// TIA Portal project "SMS-ENLAB-01-003-1501-001-PLC_V13_SP1_2_V17" (V17) (continued)
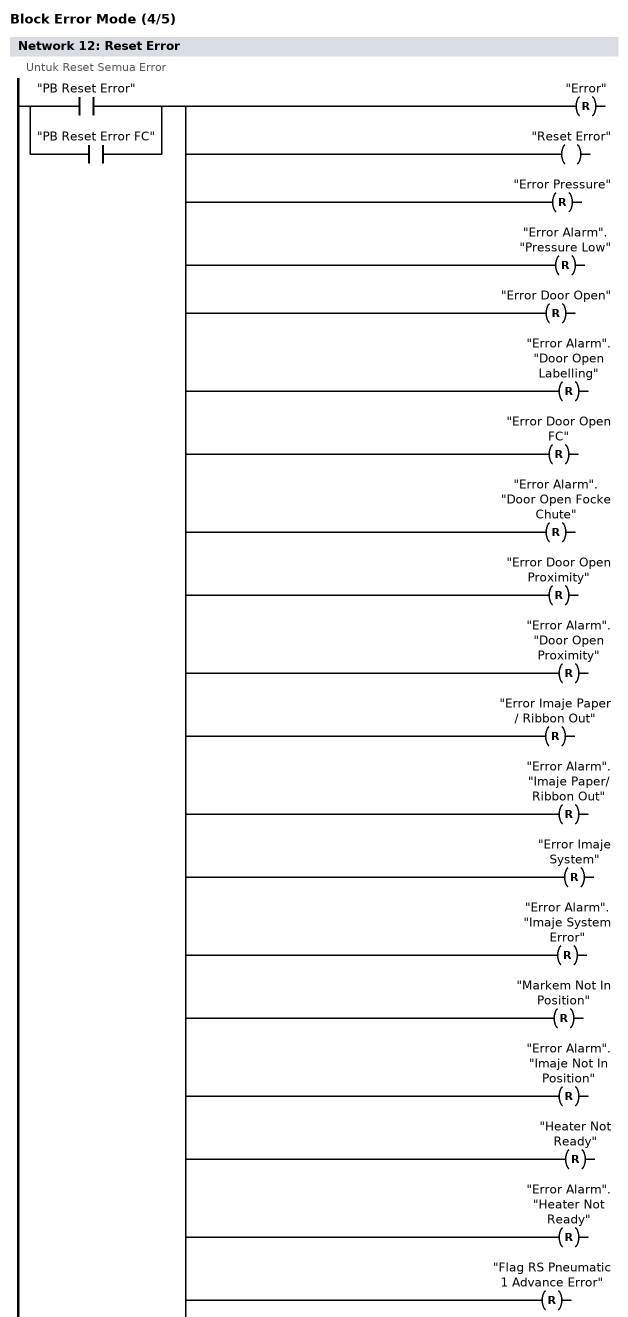
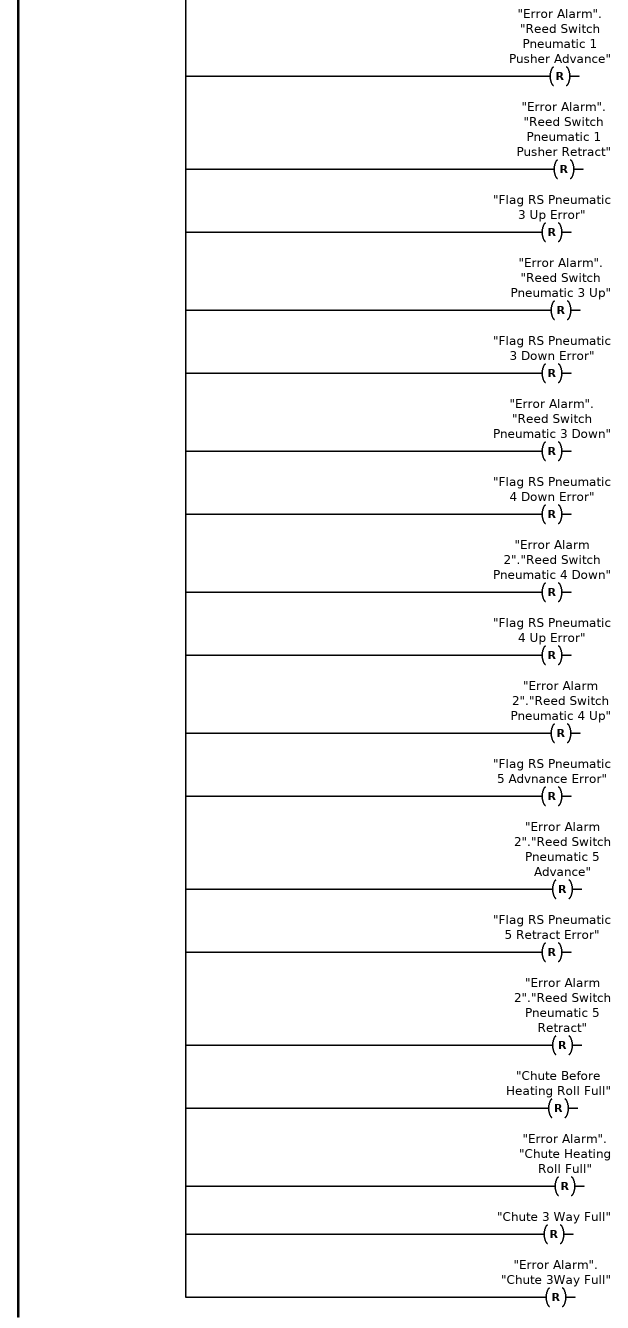
   RUNG wire#powerrail
      Contact( "PB Reset Error" )
      wire#w1
      R_Coil( "Error" )
   END_RUNG
   RUNG wire#powerrail
      Contact( "PB Reset Error FC" )
   END_RUNG wire#w1
   RUNG wire#w1
      Coil( "Reset Error" )
   END_RUNG
   RUNG wire#w1
      R_Coil( "Error Pressure" )
   END_RUNG
   RUNG wire#w1
      R_Coil( "Error Alarm"."Pressure Low" )
   END_RUNG
   RUNG wire#w1
      R_Coil( "Error Door Open" )
   END_RUNG
   RUNG wire#w1
      R_Coil( "Error Alarm"."Door Open Labelling" )
   END_RUNG
   RUNG wire#w1
      R_Coil( "Error Door Open FC" )
   END_RUNG
   RUNG wire#w1
      R_Coil( "Error Alarm"."Door Open Focke Chute" )
   END_RUNG
   RUNG wire#w1
      R_Coil( "Error Door Open Proximity" )
   END_RUNG
   RUNG wire#w1
      R_Coil( "Error Alarm"."Door Open Proximity" )
   END_RUNG
   RUNG wire#w1
      R_Coil( "Error Imaje Paper / Ribbon Out" )
   END_RUNG
   RUNG wire#w1
      R_Coil( "Error Alarm"."Imaje Paper/Ribbon Out" )
   END_RUNG
   RUNG wire#w1
      R_Coil( "Error Imaje System" )
   END_RUNG
   RUNG wire#w1
      R_Coil( "Error Alarm"."Imaje System Error" )
   END_RUNG
   RUNG wire#w1
      R_Coil( "Markem Not In Position" )
   END_RUNG
   RUNG wire#w1
      R_Coil( "Error Alarm"."Imaje Not In Position" )
   END_RUNG
   RUNG wire#w1
      R_Coil( "Heater Not Ready" )
   END_RUNG
   RUNG wire#w1
      R_Coil( "Error Alarm"."Heater Not Ready" )
   END_RUNG
   RUNG wire#w1
      R_Coil( "Flag RS Pneumatic 1 Advance Error" )
   END_RUNG
   RUNG wire#w1
      R_Coil( "Error Alarm"."Reed Switch Pneumatic 1 Pusher Advance" )
   END_RUNG
   RUNG wire#w1
      R_Coil( "Error Alarm"."Reed Switch Pneumatic 1 Pusher Retract" )
   END_RUNG
   RUNG wire#w1
      R_Coil( "Flag RS Pneumatic 3 Up Error" )
   END_RUNG
   RUNG wire#w1
      R_Coil( "Error Alarm"."Reed Switch Pneumatic 3 Up" )
   END_RUNG
   RUNG wire#w1
      R_Coil( "Flag RS Pneumatic 3 Down Error" )
   END_RUNG
   RUNG wire#w1
      R_Coil( "Error Alarm"."Reed Switch Pneumatic 3 Down" )
   END_RUNG
   RUNG wire#w1
      R_Coil( "Flag RS Pneumatic 4 Down Error" )
   END_RUNG
   RUNG wire#w1
      R_Coil( "Error Alarm 2"."Reed Switch Pneumatic 4 Down" )
   END_RUNG
   RUNG wire#w1
      R_Coil( "Flag RS Pneumatic 4 Up Error" )
   END_RUNG
   RUNG wire#w1
      R_Coil( "Error Alarm 2"."Reed Switch Pneumatic 4 Up" )
   END_RUNG
   RUNG wire#w1
      R_Coil( "Flag RS Pneumatic 5 Advnance Error" )
   END_RUNG
   RUNG wire#w1
      R_Coil( "Error Alarm 2"."Reed Switch Pneumatic 5 Advance" )
   END_RUNG
   RUNG wire#w1
      R_Coil( "Flag RS Pneumatic 5 Retract Error" )
   END_RUNG
   RUNG wire#w1
      R_Coil( "Error Alarm 2"."Reed Switch Pneumatic 5 Retract" )
   END_RUNG
   RUNG wire#w1
      R_Coil( "Chute Before Heating Roll Full" )
   END_RUNG
   RUNG wire#w1
      R_Coil( "Error Alarm"."Chute Heating Roll Full" )
   END_RUNG
   RUNG wire#w1
      R_Coil( "Chute 3 Way Full" )
   END_RUNG
   RUNG wire#w1
      R_Coil( "Error Alarm"."Chute 3Way Full" )
   END_RUNG
   // the same network as SCL:
   #_w1 := "PB Reset Error" OR "PB Reset Error FC";
   IF #_w1 THEN "Error" := FALSE; END_IF;
   "Reset Error" := #_w1;
   IF #_w1 THEN
       "Error Pressure" := FALSE;
       "Error Alarm"."Pressure Low" := FALSE;
       "Error Door Open" := FALSE;
       "Error Alarm"."Door Open Labelling" := FALSE;
       "Error Door Open FC" := FALSE;
       "Error Alarm"."Door Open Focke Chute" := FALSE;
       "Error Door Open Proximity" := FALSE;
       "Error Alarm"."Door Open Proximity" := FALSE;
       "Error Imaje Paper / Ribbon Out" := FALSE;
       "Error Alarm"."Imaje Paper/Ribbon Out" := FALSE;
       "Error Imaje System" := FALSE;
       "Error Alarm"."Imaje System Error" := FALSE;
       "Markem Not In Position" := FALSE;
       "Error Alarm"."Imaje Not In Position" := FALSE;
       "Heater Not Ready" := FALSE;
       "Error Alarm"."Heater Not Ready" := FALSE;
       "Flag RS Pneumatic 1 Advance Error" := FALSE;
       "Error Alarm"."Reed Switch Pneumatic 1 Pusher Advance" := FALSE;
       "Error Alarm"."Reed Switch Pneumatic 1 Pusher Retract" := FALSE;
       "Flag RS Pneumatic 3 Up Error" := FALSE;
       "Error Alarm"."Reed Switch Pneumatic 3 Up" := FALSE;
       "Flag RS Pneumatic 3 Down Error" := FALSE;
       "Error Alarm"."Reed Switch Pneumatic 3 Down" := FALSE;
       "Flag RS Pneumatic 4 Down Error" := FALSE;
       "Error Alarm 2"."Reed Switch Pneumatic 4 Down" := FALSE;
       "Flag RS Pneumatic 4 Up Error" := FALSE;
       "Error Alarm 2"."Reed Switch Pneumatic 4 Up" := FALSE;
       "Flag RS Pneumatic 5 Advnance Error" := FALSE;
       "Error Alarm 2"."Reed Switch Pneumatic 5 Advance" := FALSE;
       "Flag RS Pneumatic 5 Retract Error" := FALSE;
       "Error Alarm 2"."Reed Switch Pneumatic 5 Retract" := FALSE;
       "Chute Before Heating Roll Full" := FALSE;
       "Error Alarm"."Chute Heating Roll Full" := FALSE;
       "Chute 3 Way Full" := FALSE;
       "Error Alarm"."Chute 3Way Full" := FALSE;
   END_IF;
END_REGION

REGION Network 13: Enable Flow to Reject
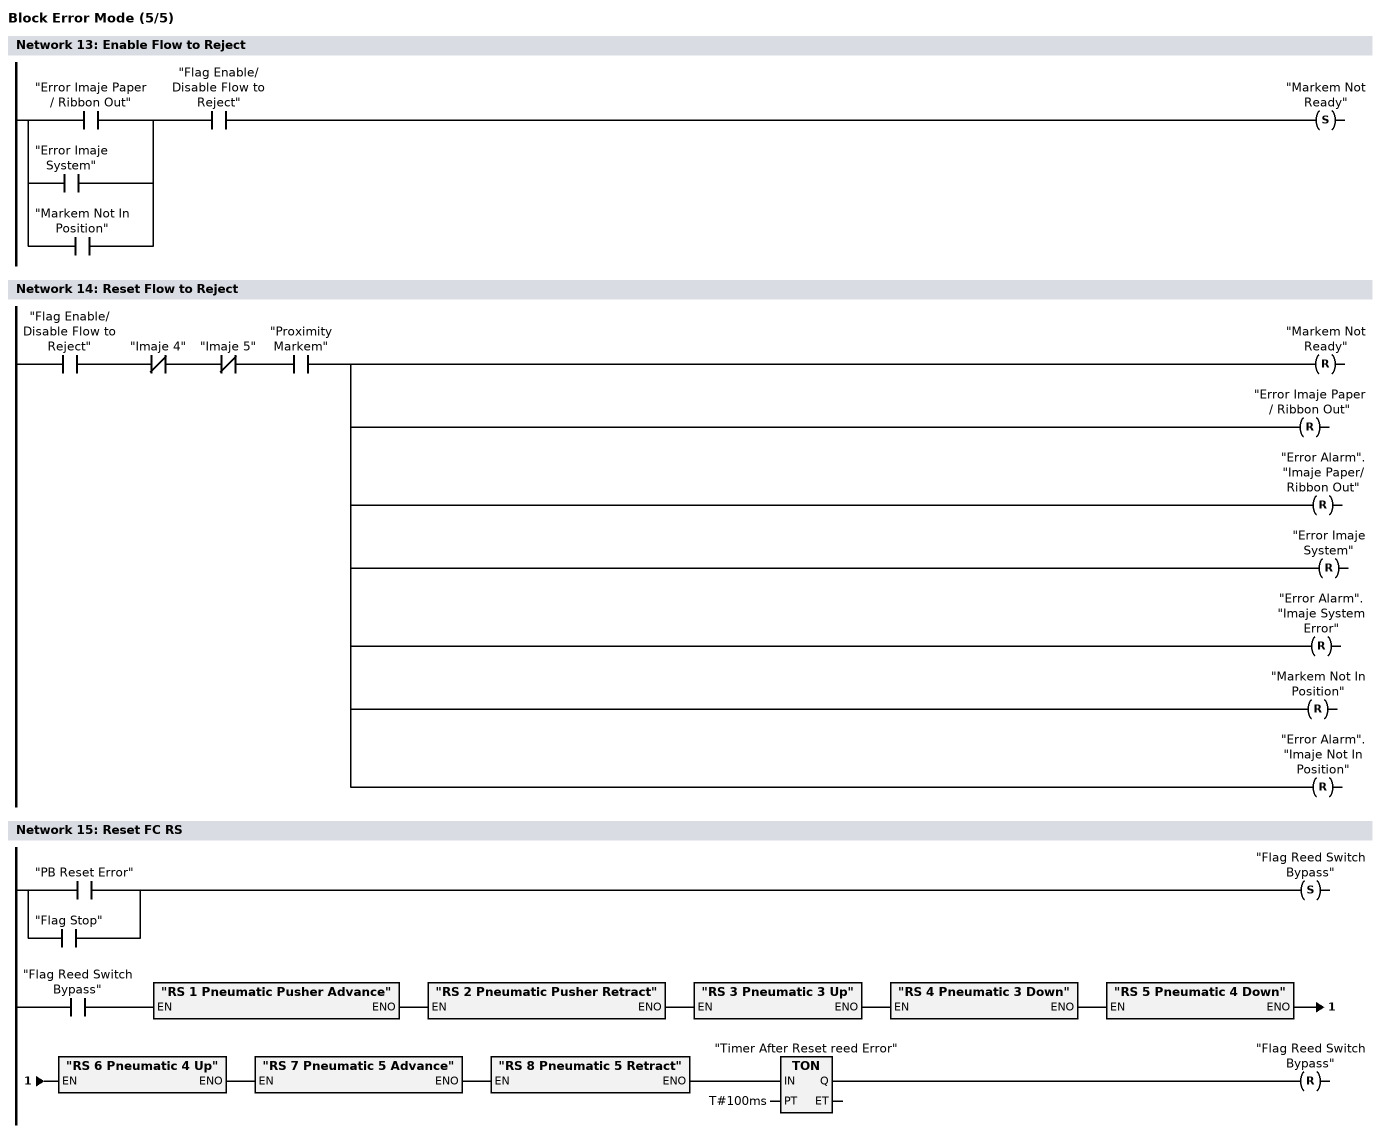
   RUNG wire#powerrail
      Contact( "Error Imaje Paper / Ribbon Out" )
      wire#w1
      Contact( "Flag Enable/Disable Flow to Reject" )
      S_Coil( "Markem Not Ready" )
   END_RUNG
   RUNG wire#powerrail
      Contact( "Error Imaje System" )
   END_RUNG wire#w1
   RUNG wire#powerrail
      Contact( "Markem Not In Position" )
   END_RUNG wire#w1
   // the same network as SCL:
   IF ("Error Imaje Paper / Ribbon Out" OR "Error Imaje System" OR "Markem Not In Position") AND "Flag Enable/Disable Flow to Reject" THEN
       "Markem Not Ready" := TRUE;
   END_IF;
END_REGION

REGION Network 14: Reset Flow to Reject
   RUNG wire#powerrail
      Contact( "Flag Enable/Disable Flow to Reject" )
      I_Contact( "Imaje 4" )
      I_Contact( "Imaje 5" )
      Contact( "Proximity Markem" )
      wire#w1
      R_Coil( "Markem Not Ready" )
   END_RUNG
   RUNG wire#w1
      R_Coil( "Error Imaje Paper / Ribbon Out" )
   END_RUNG
   RUNG wire#w1
      R_Coil( "Error Alarm"."Imaje Paper/Ribbon Out" )
   END_RUNG
   RUNG wire#w1
      R_Coil( "Error Imaje System" )
   END_RUNG
   RUNG wire#w1
      R_Coil( "Error Alarm"."Imaje System Error" )
   END_RUNG
   RUNG wire#w1
      R_Coil( "Markem Not In Position" )
   END_RUNG
   RUNG wire#w1
      R_Coil( "Error Alarm"."Imaje Not In Position" )
   END_RUNG
   // the same network as SCL:
   IF "Flag Enable/Disable Flow to Reject" AND NOT "Imaje 4" AND NOT "Imaje 5" AND "Proximity Markem" THEN
       "Markem Not Ready" := FALSE;
       "Error Imaje Paper / Ribbon Out" := FALSE;
       "Error Alarm"."Imaje Paper/Ribbon Out" := FALSE;
       "Error Imaje System" := FALSE;
       "Error Alarm"."Imaje System Error" := FALSE;
       "Markem Not In Position" := FALSE;
       "Error Alarm"."Imaje Not In Position" := FALSE;
   END_IF;
END_REGION

REGION Network 15: Reset FC RS
   IF "PB Reset Error" OR "Flag Stop" THEN "Flag Reed Switch Bypass" := TRUE; END_IF;
   "RS 1 Pneumatic Pusher Advance"(EN := "Flag Reed Switch Bypass", ENO => #_w1);
   "RS 2 Pneumatic Pusher Retract"(EN := #_w1, ENO => #_w2);
   "RS 3 Pneumatic 3 Up"(EN := #_w2, ENO => #_w3);
   "RS 4 Pneumatic 3 Down"(EN := #_w3, ENO => #_w4);
   "RS 5 Pneumatic 4 Down"(EN := #_w4, ENO => #_w5);
   "RS 6 Pneumatic 4 Up"(EN := #_w5, ENO => #_w6);
   "RS 7 Pneumatic 5 Advance"(EN := #_w6, ENO => #_w7);
   "RS 8 Pneumatic 5 Retract"(EN := #_w7, ENO => #_w8);
   "Timer After Reset reed Error".TON(IN := #_w8, PT := T#100ms);
   IF "Timer After Reset reed Error".Q THEN "Flag Reed Switch Bypass" := FALSE; END_IF;
END_REGION
END_FUNCTION_BLOCK

FUNCTION_BLOCK "Block Test Mode"   // FB2, LAD
{ S7_Optimized_Access := 'TRUE' }
VERSION : 0.1
BEGIN

REGION Network 1: Set Motor Conveyor
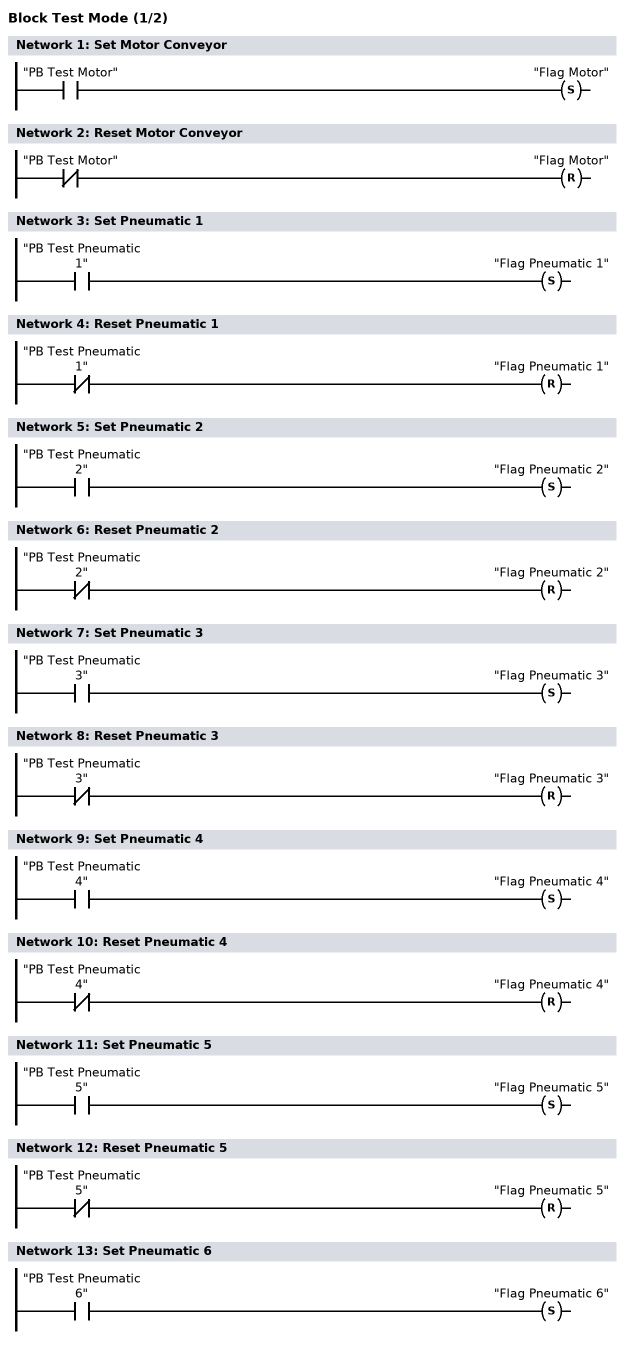
   RUNG wire#powerrail
      Contact( "PB Test Motor" )
      S_Coil( "Flag Motor" )
   END_RUNG
   // the same network as SCL:
   IF "PB Test Motor" THEN "Flag Motor" := TRUE; END_IF;
END_REGION

REGION Network 2: Reset Motor Conveyor
   RUNG wire#powerrail
      I_Contact( "PB Test Motor" )
      R_Coil( "Flag Motor" )
   END_RUNG
   // the same network as SCL:
   IF NOT "PB Test Motor" THEN "Flag Motor" := FALSE; END_IF;
END_REGION

REGION Network 3: Set Pneumatic 1
   RUNG wire#powerrail
      Contact( "PB Test Pneumatic 1" )
      S_Coil( "Flag Pneumatic 1" )
   END_RUNG
   // the same network as SCL:
   IF "PB Test Pneumatic 1" THEN "Flag Pneumatic 1" := TRUE; END_IF;
END_REGION

REGION Network 4: Reset Pneumatic 1
   RUNG wire#powerrail
      I_Contact( "PB Test Pneumatic 1" )
      R_Coil( "Flag Pneumatic 1" )
   END_RUNG
   // the same network as SCL:
   IF NOT "PB Test Pneumatic 1" THEN "Flag Pneumatic 1" := FALSE; END_IF;
END_REGION

REGION Network 5: Set Pneumatic 2
   RUNG wire#powerrail
      Contact( "PB Test Pneumatic 2" )
      S_Coil( "Flag Pneumatic 2" )
   END_RUNG
   // the same network as SCL:
   IF "PB Test Pneumatic 2" THEN "Flag Pneumatic 2" := TRUE; END_IF;
END_REGION

REGION Network 6: Reset Pneumatic 2
   RUNG wire#powerrail
      I_Contact( "PB Test Pneumatic 2" )
      R_Coil( "Flag Pneumatic 2" )
   END_RUNG
   // the same network as SCL:
   IF NOT "PB Test Pneumatic 2" THEN "Flag Pneumatic 2" := FALSE; END_IF;
END_REGION

REGION Network 7: Set Pneumatic 3
   RUNG wire#powerrail
      Contact( "PB Test Pneumatic 3" )
      S_Coil( "Flag Pneumatic 3" )
   END_RUNG
   // the same network as SCL:
   IF "PB Test Pneumatic 3" THEN "Flag Pneumatic 3" := TRUE; END_IF;
END_REGION

REGION Network 8: Reset Pneumatic 3
   RUNG wire#powerrail
      I_Contact( "PB Test Pneumatic 3" )
      R_Coil( "Flag Pneumatic 3" )
   END_RUNG
   // the same network as SCL:
   IF NOT "PB Test Pneumatic 3" THEN "Flag Pneumatic 3" := FALSE; END_IF;
END_REGION

REGION Network 9: Set Pneumatic 4
   RUNG wire#powerrail
      Contact( "PB Test Pneumatic 4" )
      S_Coil( "Flag Pneumatic 4" )
   END_RUNG
   // the same network as SCL:
   IF "PB Test Pneumatic 4" THEN "Flag Pneumatic 4" := TRUE; END_IF;
END_REGION

REGION Network 10: Reset Pneumatic 4
   RUNG wire#powerrail
      I_Contact( "PB Test Pneumatic 4" )
      R_Coil( "Flag Pneumatic 4" )
   END_RUNG
   // the same network as SCL:
   IF NOT "PB Test Pneumatic 4" THEN "Flag Pneumatic 4" := FALSE; END_IF;
END_REGION

REGION Network 11: Set Pneumatic 5
   RUNG wire#powerrail
      Contact( "PB Test Pneumatic 5" )
      S_Coil( "Flag Pneumatic 5" )
   END_RUNG
   // the same network as SCL:
   IF "PB Test Pneumatic 5" THEN "Flag Pneumatic 5" := TRUE; END_IF;
END_REGION

REGION Network 12: Reset Pneumatic 5
   RUNG wire#powerrail
      I_Contact( "PB Test Pneumatic 5" )
      R_Coil( "Flag Pneumatic 5" )
   END_RUNG
   // the same network as SCL:
   IF NOT "PB Test Pneumatic 5" THEN "Flag Pneumatic 5" := FALSE; END_IF;
END_REGION

REGION Network 13: Set Pneumatic 6
   RUNG wire#powerrail
      Contact( "PB Test Pneumatic 6" )
      S_Coil( "Flag Pneumatic 6" )
   END_RUNG
   // the same network as SCL:
   IF "PB Test Pneumatic 6" THEN "Flag Pneumatic 6" := TRUE; END_IF;
END_REGION

REGION Network 14: Reset Pneumatic 6
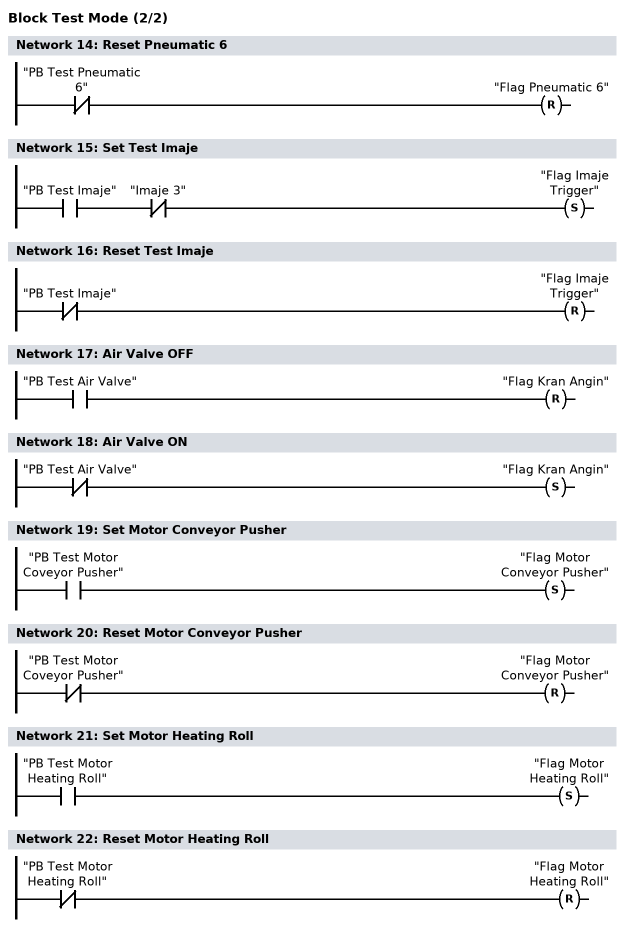
   RUNG wire#powerrail
      I_Contact( "PB Test Pneumatic 6" )
      R_Coil( "Flag Pneumatic 6" )
   END_RUNG
   // the same network as SCL:
   IF NOT "PB Test Pneumatic 6" THEN "Flag Pneumatic 6" := FALSE; END_IF;
END_REGION

REGION Network 15: Set Test Imaje
   RUNG wire#powerrail
      Contact( "PB Test Imaje" )
      I_Contact( "Imaje 3" )
      S_Coil( "Flag Imaje Trigger" )
   END_RUNG
   // the same network as SCL:
   IF "PB Test Imaje" AND NOT "Imaje 3" THEN "Flag Imaje Trigger" := TRUE; END_IF;
END_REGION

REGION Network 16: Reset Test Imaje
   RUNG wire#powerrail
      I_Contact( "PB Test Imaje" )
      R_Coil( "Flag Imaje Trigger" )
   END_RUNG
   // the same network as SCL:
   IF NOT "PB Test Imaje" THEN "Flag Imaje Trigger" := FALSE; END_IF;
END_REGION

REGION Network 17: Air Valve OFF
   RUNG wire#powerrail
      Contact( "PB Test Air Valve" )
      R_Coil( "Flag Kran Angin" )
   END_RUNG
   // the same network as SCL:
   IF "PB Test Air Valve" THEN "Flag Kran Angin" := FALSE; END_IF;
END_REGION

REGION Network 18: Air Valve ON
   RUNG wire#powerrail
      I_Contact( "PB Test Air Valve" )
      S_Coil( "Flag Kran Angin" )
   END_RUNG
   // the same network as SCL:
   IF NOT "PB Test Air Valve" THEN "Flag Kran Angin" := TRUE; END_IF;
END_REGION

REGION Network 19: Set Motor Conveyor Pusher
   RUNG wire#powerrail
      Contact( "PB Test Motor Coveyor Pusher" )
      S_Coil( "Flag Motor Conveyor Pusher" )
   END_RUNG
   // the same network as SCL:
   IF "PB Test Motor Coveyor Pusher" THEN "Flag Motor Conveyor Pusher" := TRUE; END_IF;
END_REGION

REGION Network 20: Reset Motor Conveyor Pusher
   RUNG wire#powerrail
      I_Contact( "PB Test Motor Coveyor Pusher" )
      R_Coil( "Flag Motor Conveyor Pusher" )
   END_RUNG
   // the same network as SCL:
   IF NOT "PB Test Motor Coveyor Pusher" THEN "Flag Motor Conveyor Pusher" := FALSE; END_IF;
END_REGION

REGION Network 21: Set Motor Heating Roll
   RUNG wire#powerrail
      Contact( "PB Test Motor Heating Roll" )
      S_Coil( "Flag Motor Heating Roll" )
   END_RUNG
   // the same network as SCL:
   IF "PB Test Motor Heating Roll" THEN "Flag Motor Heating Roll" := TRUE; END_IF;
END_REGION

REGION Network 22: Reset Motor Heating Roll
   RUNG wire#powerrail
      I_Contact( "PB Test Motor Heating Roll" )
      R_Coil( "Flag Motor Heating Roll" )
   END_RUNG
   // the same network as SCL:
   IF NOT "PB Test Motor Heating Roll" THEN "Flag Motor Heating Roll" := FALSE; END_IF;
END_REGION
END_FUNCTION_BLOCK

FUNCTION_BLOCK "Block Output"   // FB3, LAD
{ S7_Optimized_Access := 'TRUE' }
VERSION : 0.1
BEGIN

REGION Network 1: Red Light Tower
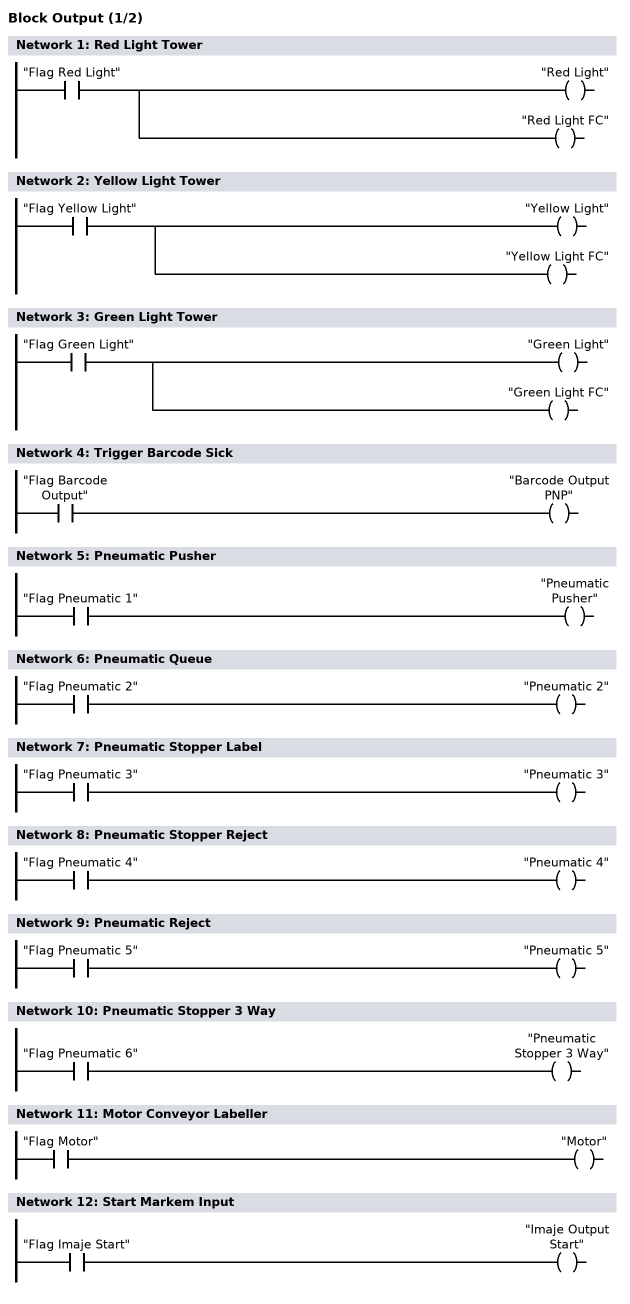
   RUNG wire#powerrail
      Contact( "Flag Red Light" )
      wire#w1
      Coil( "Red Light" )
   END_RUNG
   RUNG wire#w1
      Coil( "Red Light FC" )
   END_RUNG
   // the same network as SCL:
   "Red Light" := "Flag Red Light";
   "Red Light FC" := "Flag Red Light";
END_REGION

REGION Network 2: Yellow Light Tower
   RUNG wire#powerrail
      Contact( "Flag Yellow Light" )
      wire#w1
      Coil( "Yellow Light" )
   END_RUNG
   RUNG wire#w1
      Coil( "Yellow Light FC" )
   END_RUNG
   // the same network as SCL:
   "Yellow Light" := "Flag Yellow Light";
   "Yellow Light FC" := "Flag Yellow Light";
END_REGION

REGION Network 3: Green Light Tower
   RUNG wire#powerrail
      Contact( "Flag Green Light" )
      wire#w1
      Coil( "Green Light" )
   END_RUNG
   RUNG wire#w1
      Coil( "Green Light FC" )
   END_RUNG
   // the same network as SCL:
   "Green Light" := "Flag Green Light";
   "Green Light FC" := "Flag Green Light";
END_REGION

REGION Network 4: Trigger Barcode Sick
   RUNG wire#powerrail
      Contact( "Flag Barcode Output" )
      Coil( "Barcode Output PNP" )
   END_RUNG
   // the same network as SCL:
   "Barcode Output PNP" := "Flag Barcode Output";
END_REGION

REGION Network 5: Pneumatic Pusher
   RUNG wire#powerrail
      Contact( "Flag Pneumatic 1" )
      Coil( "Pneumatic Pusher" )
   END_RUNG
   // the same network as SCL:
   "Pneumatic Pusher" := "Flag Pneumatic 1";
END_REGION

REGION Network 6: Pneumatic Queue
   RUNG wire#powerrail
      Contact( "Flag Pneumatic 2" )
      Coil( "Pneumatic 2" )
   END_RUNG
   // the same network as SCL:
   "Pneumatic 2" := "Flag Pneumatic 2";
END_REGION

REGION Network 7: Pneumatic Stopper Label
   RUNG wire#powerrail
      Contact( "Flag Pneumatic 3" )
      Coil( "Pneumatic 3" )
   END_RUNG
   // the same network as SCL:
   "Pneumatic 3" := "Flag Pneumatic 3";
END_REGION

REGION Network 8: Pneumatic Stopper Reject
   RUNG wire#powerrail
      Contact( "Flag Pneumatic 4" )
      Coil( "Pneumatic 4" )
   END_RUNG
   // the same network as SCL:
   "Pneumatic 4" := "Flag Pneumatic 4";
END_REGION

REGION Network 9: Pneumatic Reject
   RUNG wire#powerrail
      Contact( "Flag Pneumatic 5" )
      Coil( "Pneumatic 5" )
   END_RUNG
   // the same network as SCL:
   "Pneumatic 5" := "Flag Pneumatic 5";
END_REGION

REGION Network 10: Pneumatic Stopper 3 Way
   RUNG wire#powerrail
      Contact( "Flag Pneumatic 6" )
      Coil( "Pneumatic Stopper 3 Way" )
   END_RUNG
   // the same network as SCL:
   "Pneumatic Stopper 3 Way" := "Flag Pneumatic 6";
END_REGION

REGION Network 11: Motor Conveyor Labeller
   RUNG wire#powerrail
      Contact( "Flag Motor" )
      Coil( "Motor" )
   END_RUNG
   // the same network as SCL:
   "Motor" := "Flag Motor";
END_REGION

REGION Network 12: Start Markem Input
   RUNG wire#powerrail
      Contact( "Flag Imaje Start" )
      Coil( "Imaje Output Start" )
   END_RUNG
   // the same network as SCL:
   "Imaje Output Start" := "Flag Imaje Start";
END_REGION

REGION Network 13: Pause Markem Input
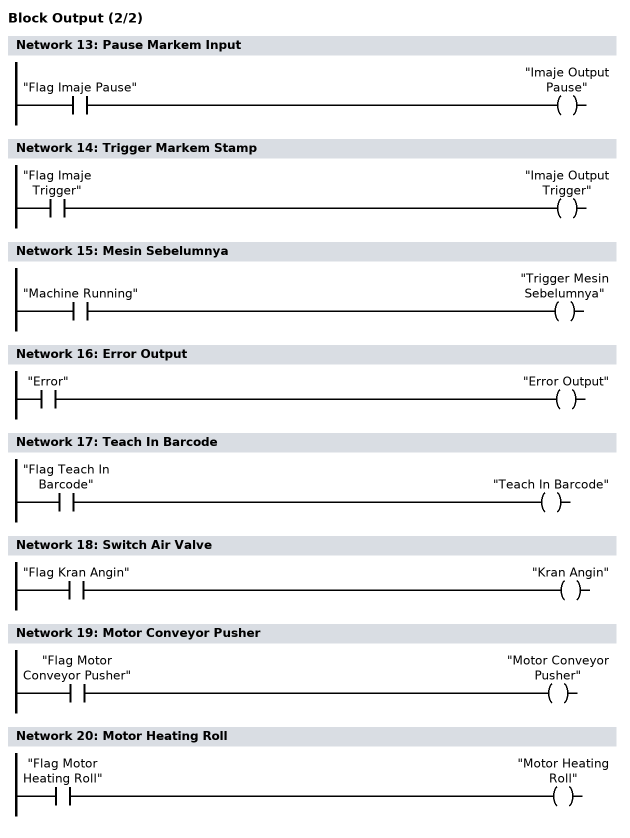
   RUNG wire#powerrail
      Contact( "Flag Imaje Pause" )
      Coil( "Imaje Output Pause" )
   END_RUNG
   // the same network as SCL:
   "Imaje Output Pause" := "Flag Imaje Pause";
END_REGION

REGION Network 14: Trigger Markem Stamp
   RUNG wire#powerrail
      Contact( "Flag Imaje Trigger" )
      Coil( "Imaje Output Trigger" )
   END_RUNG
   // the same network as SCL:
   "Imaje Output Trigger" := "Flag Imaje Trigger";
END_REGION

REGION Network 15: Mesin Sebelumnya
   RUNG wire#powerrail
      Contact( "Machine Running" )
      Coil( "Trigger Mesin Sebelumnya" )
   END_RUNG
   // the same network as SCL:
   "Trigger Mesin Sebelumnya" := "Machine Running";
END_REGION

REGION Network 16: Error Output
   RUNG wire#powerrail
      Contact( "Error" )
      Coil( "Error Output" )
   END_RUNG
   // the same network as SCL:
   "Error Output" := "Error";
END_REGION

REGION Network 17: Teach In Barcode
   RUNG wire#powerrail
      Contact( "Flag Teach In Barcode" )
      Coil( "Teach In Barcode" )
   END_RUNG
   // the same network as SCL:
   "Teach In Barcode" := "Flag Teach In Barcode";
END_REGION

REGION Network 18: Switch Air Valve
   RUNG wire#powerrail
      Contact( "Flag Kran Angin" )
      Coil( "Kran Angin" )
   END_RUNG
   // the same network as SCL:
   "Kran Angin" := "Flag Kran Angin";
END_REGION

REGION Network 19: Motor Conveyor Pusher
   RUNG wire#powerrail
      Contact( "Flag Motor Conveyor Pusher" )
      Coil( "Motor Conveyor Pusher" )
   END_RUNG
   // the same network as SCL:
   "Motor Conveyor Pusher" := "Flag Motor Conveyor Pusher";
END_REGION

REGION Network 20: Motor Heating Roll
   RUNG wire#powerrail
      Contact( "Flag Motor Heating Roll" )
      Coil( "Motor Heating Roll" )
   END_RUNG
   // the same network as SCL:
   "Motor Heating Roll" := "Flag Motor Heating Roll";
END_REGION
END_FUNCTION_BLOCK

FUNCTION_BLOCK "S Block Current Shift"   // FB4, LAD
{ S7_Optimized_Access := 'TRUE' }
VERSION : 0.1
   VAR_TEMP   // added for the SCL form of the ladder/FBD networks
      _w1 : Bool;
   END_VAR
BEGIN

REGION Network 1: Input Sloft
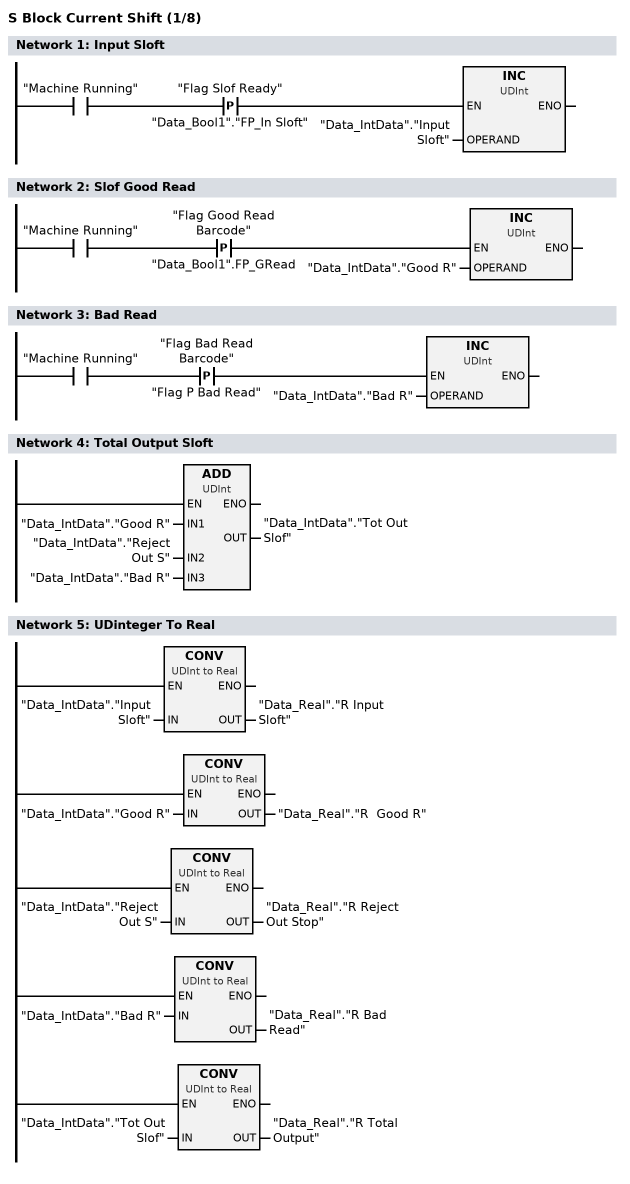
   RUNG wire#powerrail
      Contact( "Machine Running" )
      P_Contact(operand := "Flag Slof Ready", bit := "Data_Bool1"."FP_In Sloft")
      { S7_Templates := "DestType := UDInt"; S7_GenerateENO := "TRUE" } Inc( "Data_IntData"."Input Sloft" )
   END_RUNG
   // the same network as SCL:
   #_w1 := "Machine Running" AND "Flag Slof Ready" AND NOT "Data_Bool1"."FP_In Sloft";   // rising edge of "Flag Slof Ready"
   "Data_Bool1"."FP_In Sloft" := "Flag Slof Ready";
   IF #_w1 THEN "Data_IntData"."Input Sloft" := "Data_IntData"."Input Sloft" + 1; END_IF;
END_REGION

REGION Network 2: Slof Good Read
   RUNG wire#powerrail
      Contact( "Machine Running" )
      P_Contact(operand := "Flag Good Read Barcode", bit := "Data_Bool1".FP_GRead)
      { S7_Templates := "DestType := UDInt"; S7_GenerateENO := "TRUE" } Inc( "Data_IntData"."Good R" )
   END_RUNG
   // the same network as SCL:
   #_w1 := "Machine Running" AND "Flag Good Read Barcode" AND NOT "Data_Bool1".FP_GRead;   // rising edge of "Flag Good Read Barcode"
   "Data_Bool1".FP_GRead := "Flag Good Read Barcode";
   IF #_w1 THEN "Data_IntData"."Good R" := "Data_IntData"."Good R" + 1; END_IF;
END_REGION

REGION Network 3: Bad Read
   RUNG wire#powerrail
      Contact( "Machine Running" )
      P_Contact(operand := "Flag Bad Read Barcode", bit := "Flag P Bad Read")
      { S7_Templates := "DestType := UDInt"; S7_GenerateENO := "TRUE" } Inc( "Data_IntData"."Bad R" )
   END_RUNG
   // the same network as SCL:
   #_w1 := "Machine Running" AND "Flag Bad Read Barcode" AND NOT "Flag P Bad Read";   // rising edge of "Flag Bad Read Barcode"
   "Flag P Bad Read" := "Flag Bad Read Barcode";
   IF #_w1 THEN "Data_IntData"."Bad R" := "Data_IntData"."Bad R" + 1; END_IF;
END_REGION

REGION Network 4: Total Output Sloft
   RUNG wire#powerrail
      { S7_Templates := "SrcType := UDInt"; S7_GenerateENO := "TRUE" } Add(in1 := "Data_IntData"."Good R", in2 := "Data_IntData"."Reject Out S", in3 := "Data_IntData"."Bad R", out => "Data_IntData"."Tot Out Slof")
   END_RUNG
   // the same network as SCL:
   "Data_IntData"."Tot Out Slof" := "Data_IntData"."Good R" + "Data_IntData"."Reject Out S" + "Data_IntData"."Bad R";
END_REGION

REGION Network 5: UDinteger To Real
   RUNG wire#powerrail
      { S7_Templates := "[SrcType := UDInt, DestType := Real]"; S7_GenerateENO := "TRUE" } Convert(in := "Data_IntData"."Input Sloft", out => "Data_Real"."R Input Sloft")
   END_RUNG
   RUNG wire#powerrail
      { S7_Templates := "[SrcType := UDInt, DestType := Real]"; S7_GenerateENO := "TRUE" } Convert(in := "Data_IntData"."Good R", out => "Data_Real"."R  Good R")
   END_RUNG
   RUNG wire#powerrail
      { S7_Templates := "[SrcType := UDInt, DestType := Real]"; S7_GenerateENO := "TRUE" } Convert(in := "Data_IntData"."Reject Out S", out => "Data_Real"."R Reject Out Stop")
   END_RUNG
   RUNG wire#powerrail
      { S7_Templates := "[SrcType := UDInt, DestType := Real]"; S7_GenerateENO := "TRUE" } Convert(in := "Data_IntData"."Bad R", out => "Data_Real"."R Bad Read")
   END_RUNG
   RUNG wire#powerrail
      { S7_Templates := "[SrcType := UDInt, DestType := Real]"; S7_GenerateENO := "TRUE" } Convert(in := "Data_IntData"."Tot Out Slof", out => "Data_Real"."R Total Output")
   END_RUNG
   // the same network as SCL:
   "Data_Real"."R Input Sloft" := UDINT_TO_REAL("Data_IntData"."Input Sloft");
   "Data_Real"."R  Good R" := UDINT_TO_REAL("Data_IntData"."Good R");
   "Data_Real"."R Reject Out Stop" := UDINT_TO_REAL("Data_IntData"."Reject Out S");
   "Data_Real"."R Bad Read" := UDINT_TO_REAL("Data_IntData"."Bad R");
   "Data_Real"."R Total Output" := UDINT_TO_REAL("Data_IntData"."Tot Out Slof");
END_REGION

REGION Network 6: % Sloft terhadap Input Sloft
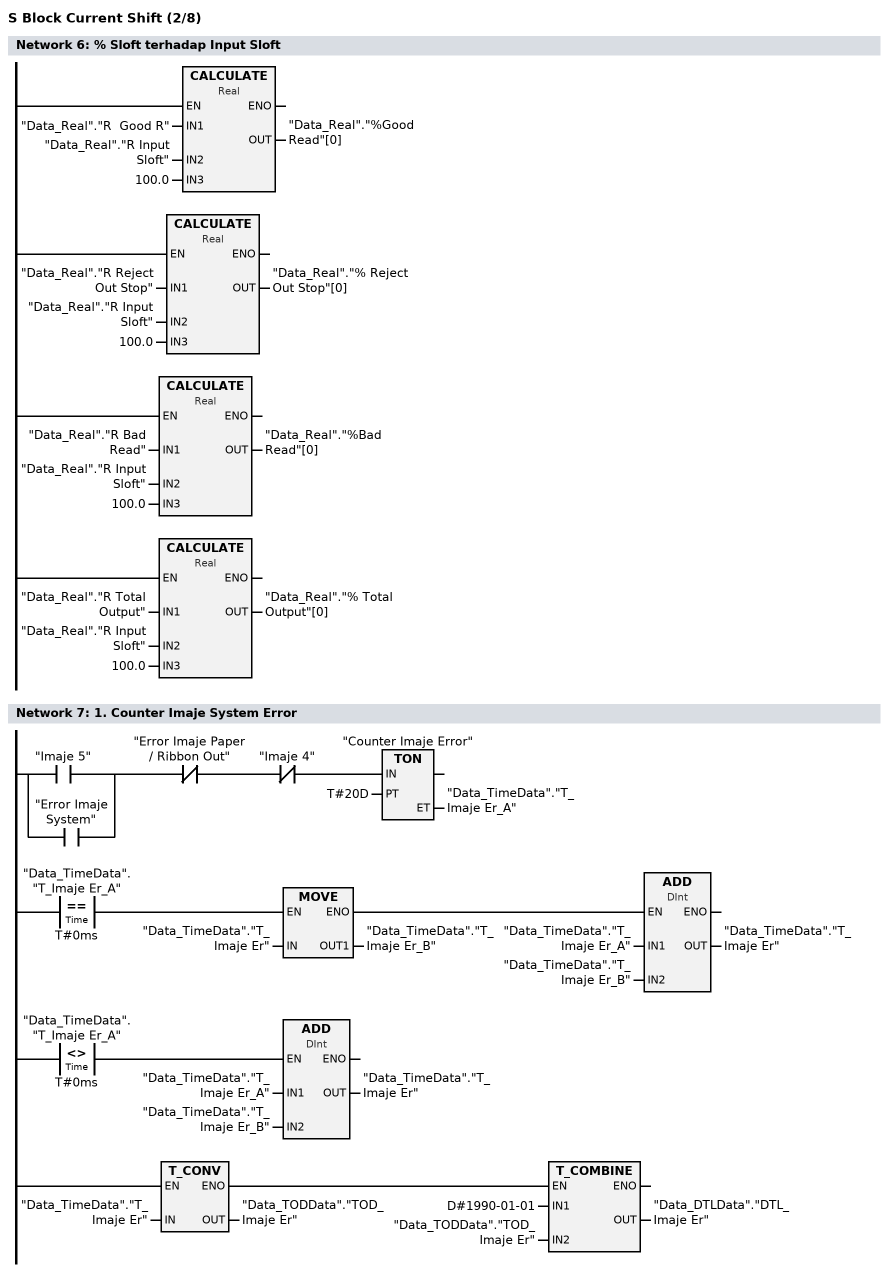
   RUNG wire#powerrail
      { S7_Templates := "SrcType := Real"; S7_GenerateENO := "TRUE"; S7_Expression := "(IN1/IN2)*IN3" } Calculate(in1 := "Data_Real"."R  Good R", in2 := "Data_Real"."R Input Sloft", in3 := 100.0, out => "Data_Real"."%Good Read"[0])
   END_RUNG
   RUNG wire#powerrail
      { S7_Templates := "SrcType := Real"; S7_GenerateENO := "TRUE"; S7_Expression := "(IN1/IN2)*IN3" } Calculate(in1 := "Data_Real"."R Reject Out Stop", in2 := "Data_Real"."R Input Sloft", in3 := 100.0, out => "Data_Real"."% Reject Out Stop"[0])
   END_RUNG
   RUNG wire#powerrail
      { S7_Templates := "SrcType := Real"; S7_GenerateENO := "TRUE"; S7_Expression := "(IN1/IN2)*IN3" } Calculate(in1 := "Data_Real"."R Bad Read", in2 := "Data_Real"."R Input Sloft", in3 := 100.0, out => "Data_Real"."%Bad Read"[0])
   END_RUNG
   RUNG wire#powerrail
      { S7_Templates := "SrcType := Real"; S7_GenerateENO := "TRUE"; S7_Expression := "(IN1/IN2)*IN3" } Calculate(in1 := "Data_Real"."R Total Output", in2 := "Data_Real"."R Input Sloft", in3 := 100.0, out => "Data_Real"."% Total Output"[0])
   END_RUNG
   // the same network as SCL:
   "Data_Real"."%Good Read"[0] := ("Data_Real"."R  Good R"/"Data_Real"."R Input Sloft")*100.0;
   "Data_Real"."% Reject Out Stop"[0] := ("Data_Real"."R Reject Out Stop"/"Data_Real"."R Input Sloft")*100.0;
   "Data_Real"."%Bad Read"[0] := ("Data_Real"."R Bad Read"/"Data_Real"."R Input Sloft")*100.0;
   "Data_Real"."% Total Output"[0] := ("Data_Real"."R Total Output"/"Data_Real"."R Input Sloft")*100.0;
END_REGION

REGION Network 7: 1. Counter Imaje System Error
   // ENO of a box is taken as its EN; it also drops when the box reports an error
   "Counter Imaje Error".TON(IN := ("Imaje 5" OR "Error Imaje System") AND NOT "Error Imaje Paper / Ribbon Out" AND NOT "Imaje 4",
                           PT := T#20D,
                           ET => "Data_TimeData"."T_Imaje Er_A");
   IF "Data_TimeData"."T_Imaje Er_A" = T#0ms THEN
       "Data_TimeData"."T_Imaje Er_B" := "Data_TimeData"."T_Imaje Er";
       "Data_TimeData"."T_Imaje Er" := "Data_TimeData"."T_Imaje Er_A" + "Data_TimeData"."T_Imaje Er_B";
   END_IF;
   IF "Data_TimeData"."T_Imaje Er_A" <> T#0ms THEN
       "Data_TimeData"."T_Imaje Er" := "Data_TimeData"."T_Imaje Er_A" + "Data_TimeData"."T_Imaje Er_B";
   END_IF;
   "Data_TODData"."TOD_Imaje Er" := T_CONV(IN := "Data_TimeData"."T_Imaje Er");
   "Data_DTLData"."DTL_Imaje Er" := T_COMBINE(IN1 := D#1990-01-01, IN2 := "Data_TODData"."TOD_Imaje Er");
END_REGION

REGION Network 8: 2. Paper Ribbon Out
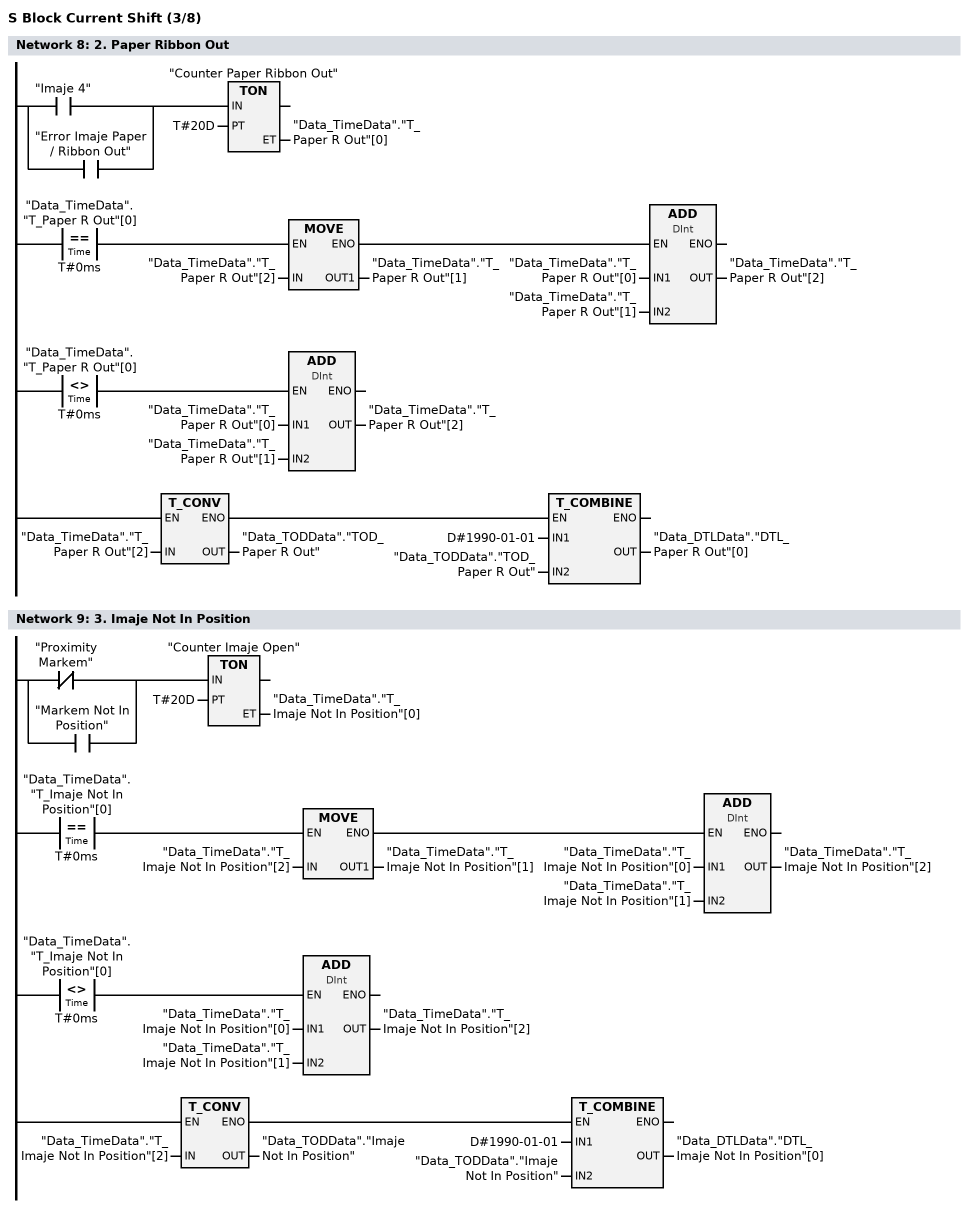
   // ENO of a box is taken as its EN; it also drops when the box reports an error
   "Counter Paper Ribbon Out".TON(IN := "Imaje 4" OR "Error Imaje Paper / Ribbon Out",
                           PT := T#20D,
                           ET => "Data_TimeData"."T_Paper R Out"[0]);
   #_w1 := "Data_TimeData"."T_Paper R Out"[0] = T#0ms;
   IF #_w1 THEN
       "Data_TimeData"."T_Paper R Out"[1] := "Data_TimeData"."T_Paper R Out"[2];
       "Data_TimeData"."T_Paper R Out"[2] := "Data_TimeData"."T_Paper R Out"[0] + "Data_TimeData"."T_Paper R Out"[1];
   END_IF;
   IF "Data_TimeData"."T_Paper R Out"[0] <> T#0ms THEN
       "Data_TimeData"."T_Paper R Out"[2] := "Data_TimeData"."T_Paper R Out"[0] + "Data_TimeData"."T_Paper R Out"[1];
   END_IF;
   "Data_TODData"."TOD_Paper R Out" := T_CONV(IN := "Data_TimeData"."T_Paper R Out"[2]);
   "Data_DTLData"."DTL_Paper R Out"[0] := T_COMBINE(IN1 := D#1990-01-01,
                           IN2 := "Data_TODData"."TOD_Paper R Out");
END_REGION

REGION Network 9: 3. Imaje Not In Position
   // ENO of a box is taken as its EN; it also drops when the box reports an error
   "Counter Imaje Open".TON(IN := NOT "Proximity Markem" OR "Markem Not In Position",
                           PT := T#20D,
                           ET => "Data_TimeData"."T_Imaje Not In Position"[0]);
   #_w1 := "Data_TimeData"."T_Imaje Not In Position"[0] = T#0ms;
   IF #_w1 THEN
       "Data_TimeData"."T_Imaje Not In Position"[1] := "Data_TimeData"."T_Imaje Not In Position"[2];
       "Data_TimeData"."T_Imaje Not In Position"[2] := "Data_TimeData"."T_Imaje Not In Position"[0] + "Data_TimeData"."T_Imaje Not In Position"[1];
   END_IF;
   IF "Data_TimeData"."T_Imaje Not In Position"[0] <> T#0ms THEN
       "Data_TimeData"."T_Imaje Not In Position"[2] := "Data_TimeData"."T_Imaje Not In Position"[0] + "Data_TimeData"."T_Imaje Not In Position"[1];
   END_IF;
   "Data_TODData"."Imaje Not In Position" := T_CONV(IN := "Data_TimeData"."T_Imaje Not In Position"[2]);
   "Data_DTLData"."DTL_Imaje Not In Position"[0] := T_COMBINE(IN1 := D#1990-01-01,
                           IN2 := "Data_TODData"."Imaje Not In Position");
END_REGION

REGION Network 10: 4. Counter Pressure Low